REGION Network 11: External containerstation
         ON    "DB702_Tank_Value".Tank[1].With_ContainerStation;
         O     "DB009_Faults".Faults_Reset_FKT_M1;
         R     "DB822_Error_Tank".InterfaceContainer.FLT_SupplyContainerstation;
         R     "DB822_Error_Tank".InterfaceContainer.FLT_containerstation;
         R     "DB822_Error_Tank".InterfaceContainer.FLT_containerNotReady_C1;
   //-----
         AN    "Container_FaultSupply";
         A     "DB702_Tank_Value".Tank[1].With_ContainerStation;
         AN    "DB822_Error_Tank".InterfaceContainer.FLT_SupplyContainerstation;
         S     "DB822_Error_Tank".InterfaceContainer.FLT_SupplyContainerstation;
         S     "DB009_Faults".Faultschanging_M1;
   //---
   //      U     "Container_Faulty"
   //      U     "DB702_Tank_Value".Tank[1].With_ContainerStation
   //      UN    "DB822_Error_Tank".InterfaceContainer.FLT_containerstation
   //      S     "DB822_Error_Tank".InterfaceContainer.FLT_containerstation
   //      S     "DB009_Faults".Faultschanging_M1
   //---
         A     "ES_Container_C1";
         A     "DB702_Tank_Value".Tank[1].With_ContainerStation;
         =     "DB822_Error_Tank".InterfaceContainer.MSG_EScontainerstation;
   //---
         AN    "Container_Ready_C1";
         A     "DB702_Tank_Value".Tank[1].With_ContainerStation;
         A     "DB612_Tank_State".Tank[1].Switch_Refilling_ON_OFF;
         A     "DB619_State_MPart".Operationmode[1].Controllvoltage;
         AN    "DB822_Error_Tank".InterfaceContainer.FLT_containerNotReady_C1;
         S     "DB822_Error_Tank".InterfaceContainer.FLT_containerNotReady_C1;
         S     "DB009_Faults".Faultschanging_M1;
   //---
         AN    "Container_Ready_C1";
         A     "DB702_Tank_Value".Tank[1].With_ContainerStation;
         A     "DB619_State_MPart".Operationmode[1].Controllvoltage;
         A     "DB612_Tank_State".Tank[1].Switch_Refilling_ON_OFF;
         AN    "DB822_Error_Tank".InterfaceContainer.FLT_containerNotReady_C1;
         =     "DB822_Error_Tank".InterfaceContainer.MSG_containerNotReady_C1;
   //---
         O     "DB822_Error_Tank".InterfaceContainer.FLT_SupplyContainerstation;
         O     "DB822_Error_Tank".InterfaceContainer.FLT_containerstation;
         O     "DB822_Error_Tank".InterfaceContainer.FLT_containerNotReady_C1;
         S     "DB009_Faults".Faults_FKT_Grp_3_M1;
   //---
END_REGION

REGION Network 12: A fault exists
         O     "DB612_Tank_State".Tank[1].Fault_Exist;
         O     "DB612_Tank_State".Agitator[1].FLT_Exist;
         O     "DB612_Tank_State".AgitatorBarell[1].FLT_Exist;
         O     "DB612_Tank_State".Vacuum[1].FLT_PVacuum;
         O     "DB612_Tank_State".CirculationPump[1].FaultExist;
         O     "DB612_Tank_State".ControllerTankTemp[1].Fault_Exist;
         O     "DB612_Tank_State".ControllerTankJacketHeater[1].Fault_Exist;
         O     "DB612_Tank_State".ControllerBarellTemp[1].Fault_Exist;
   //---
         O     "DB822_Error_Tank".InterfaceContainer.FLT_SupplyContainerstation;
         O     "DB822_Error_Tank".InterfaceContainer.FLT_containerstation;
         O     "DB822_Error_Tank".InterfaceContainer.FLT_containerNotReady_C1;
   //---
         =     "DB612_Tank_State".FaultExists[1];
END_REGION
END_FUNCTION_BLOCK

FUNCTION_BLOCK "FB102_Common_Aggregates_C2"   // FB102, STL
TITLE = Agitators,Tanks, Refilling, tempering
{ S7_Optimized_Access := 'FALSE' }
AUTHOR : KT242
VERSION : 0.1
// Common aggregates
   VAR_TEMP
      DINT_dummy : Real;
      CompUsedForShot : Array[1..16] of Bool;
      Dummy : Bool;
      MH_open : Bool;
      K_Tanklager : Bool;
      Valid : Bool;
      Temp_Vacuum_active : Bool;
      Temp_Cooling : Bool;
      Temp_Filling_Enable : Bool;
      Temp_StartExtern : Bool;
      Temp_WithFillingPump : Bool;
      Temp_FillingPumpActive : Bool;
      Temp_SwitchONTemp : Bool;
      Temp_EnableTempering : Bool;
      Temp_RequestFillAuto : Bool;
      HF_Pulse_alarm : Bool;
      Temp_RetVal_SFC14 : Word;
      Temp_RetVal_SFC15 : Word;
      Temp_SetValue_TG : Int;
      Temp_Refilling_Barrel : Bool;
      Temp_Filling_Valve : Bool;
   END_VAR
BEGIN

REGION Network 1: Toggle bit, if refilling over barrel station is activated
   // Copy Control bits for module to local area
         L;
         LAR1;
         L     "DB619_State_MPart".ShotMa[1].ShotData.Comp_at_Shot;
         L     "DB619_State_MPart".ShotMa[2].ShotData.Comp_at_Shot;
         OD;
         CAW;
         T     LW [ AR1 , P#0.0 ];

         A     "DB612_Tank_State".Tank[2].Switch_Refilling_from_Barrel_ON_OFF;
         =     #Temp_Refilling_Barrel;
END_REGION

REGION Network 2: Signal a mixinghead opens
         O     "DB619_State_MPart".Mixinghead[1].Shotcounter."01";
         O     "DB619_State_MPart".Mixinghead[1].Shotcounter."02";
         O     "DB619_State_MPart".Mixinghead[1].Shotcounter."03";
         O     "DB619_State_MPart".Mixinghead[1].Shotcounter."04";
         O     "DB619_State_MPart".Mixinghead[1].Shotcounter."05";
         O     "DB619_State_MPart".Mixinghead[1].Shotcounter."06";
         O     "DB619_State_MPart".Mixinghead[1].Shotcounter."07";
         O     "DB619_State_MPart".Mixinghead[1].Shotcounter."08";
         O     "DB619_State_MPart".Mixinghead[1].Shotcounter."09";
         O     "DB619_State_MPart".Mixinghead[1].Shotcounter."10";
         O     "DB619_State_MPart".Mixinghead[1].Shotcounter."11";
         O     "DB619_State_MPart".Mixinghead[1].Shotcounter."12";
         O     "DB619_State_MPart".Mixinghead[1].Shotcounter."13";
         O     "DB619_State_MPart".Mixinghead[1].Shotcounter."14";
         O     "DB619_State_MPart".Mixinghead[1].Shotcounter."15";
         O     "DB619_State_MPart".Mixinghead[1].Shotcounter."16";
         A     #CompUsedForShot[2];
         =     #MH_open;
END_REGION

REGION Network 3: Filling level
         CALL  "FC920_PV_Calc_Act_Value"
         ( IN_Act_Value_read := "DB702_Tank_Value".Tank[2].With_Level_Probe,
           IN_Act_Value_ext  := FALSE,
           IN_Ext_Value      := #DINT_dummy,
           IN_Read_Double    := FALSE,
           IN_FLT_Needful    := TRUE,
           IN_FLT_Reset      := "DB009_Faults".Faults_Reset_FKT_M1,
           IO_Any_ArrayPV    := "DB602_PV_Tank".Tank[2].Level,
           IO_Fault_Sensor   := "DB822_Error_Tank".Refilling_Tank[2].FLT_LevelSensor_broken_wire,
           IO_New_Fault      := "DB009_Faults".Faultschanging_M1,
           IO_FLT_Level_3    := "DB009_Faults".Faults_FKT_Grp_3_M1
         );
   //-----
         AN    "DB702_Tank_Value".Tank[2].DrainTank;
         R     "DB612_Tank_State".Tank[2].Switch_DrainTank_ON_OFF;
   //-----
         CALL  "FC104_FillingSignals"
         ( Tank_exist           := "DB702_Tank_Value".Tank[1].Existing,
           Actual_Level_Value   := "DB602_PV_Tank".Tank[2].Level.PV_ActV.Value,
           IN_With_Level_Probe  := "DB702_Tank_Value".Tank[2].With_Level_Probe,
           IN_With_Triptray     := "DB702_Tank_Value".Tank[2].With_Triptray,
           IN_FLT_Level_Probe   := "DB822_Error_Tank".Refilling_Tank[2].FLT_LevelSensor_broken_wire,
           IN_Max_Level         := "L_DT_max_C2",
           IN_Stop_Fill_Level   := "L_Tank_stop_C2",
           IN_Start_Fill_Level  := "L_Tank_start_C2",
           IN_Min_Level         := "L_Tank_min_C2",
           IN_Triptray          := "L_DripTray_C2",
           IN_DrainTank         := "DB612_Tank_State".Tank[2].Switch_DrainTank_ON_OFF,
           OUT_PreWarnMinLevel  := "DB612_Tank_State".Tank[2].PreWarning_Min_Level,
           OUT_Max_Level        := "DB612_Tank_State".Tank[2].Max_Level,
           OUT_Stop_Fill_Level  := "DB612_Tank_State".Tank[2].Stop_Level_Filling,
           OUT_Start_Fill_Level := "DB612_Tank_State".Tank[2].Start_Level_Filling,
           OUT_Min_Level        := "DB612_Tank_State".Tank[2].Min_Level,
           OUT_Enable_Agitator  := "DB612_Tank_State".Tank[2].Enable_Agitator,
           OUT_Triptray         := "DB612_Tank_State".Tank[2].LevelTriptray,
           IO_TankLevelPar      := "DB702_Tank_Value".Tank[2].TankLevel
         );
   //-----
END_REGION

REGION Network 4: GBE
   //      CALL  "FC920_PV_Calc_Act_Value"
   //         IN_Act_Value_read :="DB702_Tank_Value".Tank[2].With_Nucleation
   //         IN_Act_Value_ext  :=FALSE
   //         IN_Ext_Value      :=#DINT_dummy
   //         IN_Read_Double    :=FALSE
   //         IN_FLT_Needful    :=TRUE
   //         IN_FLT_Reset      :="DB009_Faults".Faults_Reset_FKT_M1
   //         IO_Any_ArrayPV    :="DB602_PV_Tank".Tank[2].Nucleation
   //         IO_Fault_Sensor   :="DB822_Error_Tank".Refilling_Tank[2].FLT_NucleationSensor_broken_wire
   //         IO_New_Fault      :="DB009_Faults".Faultschanging_M1
   //         IO_FLT_Level_3    :="DB009_Faults".Faults_FKT_Grp_3_M1
   //-----
   //      O     "DB009_Faults".Faults_Reset_FKT_M1
   //      O     "DB702_Tank_Value".Tank[2].With_Nucleation
   //      R     "DB822_Error_Tank".Refilling_Tank[2].FLT_supply_nucleation
   //      R     "DB822_Error_Tank".Refilling_Tank[2].FLT_nucleation
   //-
   //      UN    "F_GBE_C2"
   //      U     "DB702_Tank_Value".Tank[2].With_Nucleation
   //      UN    "DB822_Error_Tank".Refilling_Tank[2].FLT_supply_nucleation
   //      S     "DB009_Faults".Faultschanging_M1
   //      S     "DB822_Error_Tank".Refilling_Tank[2].FLT_supply_nucleation
   //-
   //      U     "F_GBE_Faulty_C2"
   //      U     "DB702_Tank_Value".Tank[2].With_Nucleation
   //      UN    "DB822_Error_Tank".Refilling_Tank[2].FLT_nucleation
   //      S     "DB009_Faults".Faultschanging_M1
   //      S     "DB822_Error_Tank".Refilling_Tank[2].FLT_nucleation
   //-
   //      O     "DB822_Error_Tank".Refilling_Tank[2].FLT_nucleation
   //      O     "DB822_Error_Tank".Refilling_Tank[2].FLT_supply_nucleation
   //      S     "DB009_Faults".Faults_FKT_Grp_3_M1
   //-----
END_REGION

REGION Network 5: Filling daytank
   ///----
         AN    "DB822_Error_Tank".FeedPump[2].FLT_Dryrunsafety;
         AN    "DB822_Error_Tank".FeedPump[2].FLT_Motorprotection;
         AN    "DB822_Error_Tank".FeedPump[2].FLT_No_Barrel;
         A(;
         ON    "DB702_Tank_Value".Tank[2].With_ContainerStation;
         O     "Container_Ready_C2";
         );
         A     "DB619_State_MPart".Operationmode[1].valid;
         =     #Temp_Filling_Enable;
   //-----
         A     "Container_Fillpump_run_C2";
         =     #Temp_FillingPumpActive;
   //-----
         A     "DB702_Tank_Value".Tank[2].With_ContainerStation;
         =     #Temp_WithFillingPump;
   //-----
         CALL  "FC102_Refilling"
         ( IN_Selected             := "DB702_Tank_Value".Tank[2].Existing,
           IN_ReleaseRefilling     := #Temp_Filling_Enable,
           IN_FillingPumpActive    := #Temp_FillingPumpActive,
           IN_WithFillingPump      := #Temp_WithFillingPump,
           IN_RecircWeekend        := "DB619_State_MPart".Recirculation[1].Weekendswitching,
           IN_FoamingCycleActive   := "DB619_State_MPart".Cycle[1].running,
           IN_PistonActive         := FALSE,
           IN_MH_is_open           := #MH_open,
           IN_ResetFault           := "DB009_Faults".Faults_Reset_FKT_M1,
           IN_MaxLevelTriptray     := "DB612_Tank_State".Tank[2].LevelTriptray,
           IN_PumpDeselected       := "DB753_MeteringPump".Pump[2].PumpDeselected,
           IN_SetAmountShots       := "DB702_Tank_Value".Tank[2].NoShotFilling,
           IN_PreAgitatingTime     := "DB702_Tank_Value".Tank[2].PreAgitatingTime,
           IN_FillingTimeContr     := "DB702_Tank_Value".Tank[2].FillingTimeControl,
           IN_TimeTillFillingStart := "DB702_Tank_Value".Tank[2].TimeToStartFilling,
           IN_Timer_Refilling      := "TM_Refilling_02",
           OUT_V_Preagitating      := #Dummy,
           OUT_V_Refilling         := #Temp_Filling_Valve,  //"V_ChargingTank_C2"
           OUT_R_Tankstorage       := #K_Tanklager,
           IO_Status               := "DB612_Tank_State".Tank[2],
           IO_NewFault             := "DB009_Faults".Faultschanging_M1,
           IO_FaultLevel_1         := "DB009_Faults".Faults_FKT_Grp_1_M1,
           IO_FaultLevel_2         := "DB009_Faults".Faults_FKT_Grp_2_M1,
           IO_FaultLevel_3         := "DB009_Faults".Faults_FKT_Grp_3_M1,
           IO_Fault                := "DB822_Error_Tank".Refilling_Tank[2]
         );
   //-----
         A     #Temp_Refilling_Barrel;
         JC    BarrelFill;
         R     "K_Filling_Tank_C2_TL";
         R     "V_ChargingTank_C2_2";

         A     #K_Tanklager;
         A     #Temp_Filling_Valve;
         =     "K_Filling_Tank_C2";
         =     "V_ChargingTank_C2";
         =     "V_Barrel_C2";
         =     "C_Start_Refill_ISO_ON";

         JU    NoBarrelFill;

   BarrelFill:R     "K_Filling_Tank_C2";
         R     "V_ChargingTank_C2";

         A     #K_Tanklager;
         A     #Temp_Filling_Valve;
         =     "K_Filling_Tank_C2_TL";
         =     "V_ChargingTank_C2_2";
         =     "V_Barrel_C2";
         =     "C_Start_Refill_ISO_ON";


   //-----
END_REGION

REGION Network 6: Agitator daytank
   //-----
   // Das Befüllen soll das Rührwerk nur im Auto ansteuern
   NoBarrelFill:A     "DB612_Tank_State".Tank[2].Fillingtime_runs;
         A     "DB619_State_MPart".Operationmode[1].Auto;
         =     #Temp_RequestFillAuto;

         CALL  "FC121_Aggitator"
         ( IN_Release               := "DB619_State_MPart".Operationmode[1].valid,
           IN_ControlVoltage        := "DB619_State_MPart".Operationmode[1].Controllvoltage,
           IN_Reset_fault           := "DB009_Faults".Faults_Reset_FKT_M1,
           IN_Request_Filling       := #Temp_RequestFillAuto,  //"DB612_Tank_State".Tank[2].Fillingtime_runs
           IN_Request_Feed          := 0,
           IN_Request_Cooling       := "DB612_Tank_State".ControllerTankTemp[2].CoolingActive,
           IN_Request_Heating       := "DB612_Tank_State".ControllerTankTemp[2].HeatingActive,
           IN_Fault_Motorprotection := "F_Agitator_C2",
           IN_FaultFreqConverter    := "F_FC_Agitator_C2",
           IN_MaxLevelTray          := "DB612_Tank_State".Tank[2].LevelTriptray,
           IN_EnableLevel           := "DB612_Tank_State".Tank[2].Enable_Agitator,
           IN_TimerDrive            := "TM1_Agitator_02",
           IN_TimerStartUpFConv     := "TM2_Agitator_02",
           IN_Values                := "DB702_Tank_Value".Tank[2].Agitator,
           OUT_MainsContactor       := "M_Agitator_C2",
           OUT_Release_FConverter   := "M_FU_Start_RW_K2",
           IO_Status                := "DB612_Tank_State".Agitator[2],
           IO_NewFault              := "DB009_Faults".Faultschanging_M1,
           IO_FaultLevel_3          := "DB009_Faults".Faults_FKT_Grp_3_M1,
           IO_Faults                := "DB822_Error_Tank".Agitator[2]
         );
   //-----
END_REGION

REGION Network 7: Tempering Tank
         A     "DB009_Faults".Faults_Reset_FKT_M1;
         R     "DB822_Error_Tank".ControllerTankTemp[2].Fuse_TemperingUnit;
   //-
         AN    "F_Temperiergeraet_C2";
         A     "DB702_Tank_Value".Tank[2].With_Tempering_TempGeraet;
         AN    "DB822_Error_Tank".ControllerTankTemp[2].Fuse_TemperingUnit;
         S     "DB009_Faults".Faultschanging_M1;
         S     "DB822_Error_Tank".ControllerTankTemp[2].Fuse_TemperingUnit;
   //-
         A     "DB822_Error_Tank".ControllerTankTemp[2].Fuse_TemperingUnit;
         S     "DB009_Faults".Faults_FKT_Grp_3_M1;
   //-
         CALL  "FC920_PV_Calc_Act_Value"
         ( IN_Act_Value_read := TRUE,
           IN_Act_Value_ext  := FALSE,
           IN_Ext_Value      := #DINT_dummy,
           IN_Read_Double    := FALSE,
           IN_FLT_Needful    := TRUE,
           IN_FLT_Reset      := "DB009_Faults".Faults_Reset_FKT_M1,
           IO_Any_ArrayPV    := "DB602_PV_Tank".Tank[2].Temp,
           IO_Fault_Sensor   := "DB822_Error_Tank".ControllerTankTemp[2].Sensor_FLT_broken_wire,
           IO_New_Fault      := "DB009_Faults".Faultschanging_M1,
           IO_FLT_Level_3    := "DB009_Faults".Faults_FKT_Grp_3_M1
         );
   //-----
         CALL  "FC916_PV_Limits"
         ( IN_Tolerance_Test     := TRUE,
           IN_Reset_Fault        := "DB009_Faults".Faults_Reset_FKT_M1,
           IO_Any_ArrayPV        := "DB602_PV_Tank".Tank[2].Temp,
           IO_Fault_Warn_upperL  := "DB822_Error_Tank".ControllerTankTemp[2].Warning_limit_plus,
           IO_Fault_Warn_lowerL  := "DB822_Error_Tank".ControllerTankTemp[2].Warning_limit_minus,
           IO_Fault_Alarm_upperL := "DB822_Error_Tank".ControllerTankTemp[2].Alarm_limit_plus,
           IO_Fault_Alarm_lowerL := "DB822_Error_Tank".ControllerTankTemp[2].Alarm_limit_minus,
           IO_New_Fault          := "DB009_Faults".Faultschanging_M1,
           IO_Fault_Level_1      := "DB009_Faults".Faults_FKT_Grp_2_M1,
           IO_Fault_Level_2      := #Dummy,  //"DB009_Faults".Faults_FKT_Grp_2_M1
           IO_Fault_Level_3      := "DB009_Faults".Faults_FKT_Grp_3_M1
         );
   //-----
   //---------------------------------------------
   //  Controller temperature tank Iso
   //---------------------------------------------
         O     "DB702_Tank_Value".Tank[2].With_Tempering_VKaltwasser;
         O     "DB702_Tank_Value".Tank[2].With_Tempering_Heizung;
         =     #Temp_EnableTempering;
   //---
         CALL  "FC105_Tempering"
         ( IN_Exist                := #Temp_EnableTempering,
           IN_Release              := "DB619_State_MPart".Operationmode[1].valid,
           IN_Stop_Tempering       := FALSE,
           IN_F_Fuse               := "F_Heating",
           IN_F_Limit              := FALSE,
           IN_FLT_Ackn             := "DB009_Faults".Faults_Reset_FKT_M1,
           IN_CoolingRequested     := TRUE,
           IN_HeatingRequested     := "DB702_Tank_Value".Tank[2].With_Tempering_Heizung,
           IN_actual_Temp          := "DB602_PV_Tank".Tank[2].Temp.PV_ActV.Value,
           IN_set_Temp             := "DB602_PV_Tank".Tank[2].Temp.PV_SetV.Value,
           Out_act_cooling         := #Temp_Cooling,
           Out_act_request_cooling := #Dummy,
           Out_act_heating         := "K_HeatingTank_C2",
           Out_act_request_heating := #Dummy,
           IO_StateCtrl1           := "DB612_Tank_State".ControllerTankTemp[2],
           IO_ValueCtrl1           := "DB702_Tank_Value".Pt2_Controller[2],
           IO_FaultsCtrl1          := "DB822_Error_Tank".ControllerTankTemp[2],
           IO_NewFault             := "DB009_Faults".Faultschanging_M1,
           IO_FaultLevel_3         := "DB009_Faults".Faults_FKT_Grp_3_M1
         );
   //-----
         A     "DB619_State_MPart".Machine[1].Metering."02";
         A     "DB702_Tank_Value".Tank[2].With_Tempering_WTRL;
         A     #Temp_Cooling;
         O(;
         A     "DB613_Komponent_State".HeatexchangerLP[2].CoolingActive;
         A     "DB619_State_MPart".Machine[1].Metering."02";
         A     "DB753_MeteringPump".Pump[2].WithLPHeatExchanger;
         );
         =     "V_Heatexchanger_C2";
   //-----
         ON    "DB619_State_MPart".Machine[1].Metering."02";
         ON    "DB702_Tank_Value".Tank[2].With_Tempering_WTRL;
         A     #Temp_Cooling;
         =     "V_Coolingwater_C2";
   //-----

   // Tempering device gets/sets temperature values with multiplier of 10.
         CALL  CONVERTTO
         ( IN      := "DB602_PV_Tank".Tank[2].Temp.PV_SetV.Value,
           Ret_Val := #Temp_SetValue_TG
         );

         L     #Temp_SetValue_TG;
         L     10;
         *I;
         T     #Temp_SetValue_TG;

         A     "Flag_00_500_Hertz";
         FP    "HF_pulse_alarm_GWK2";
         =     #HF_Pulse_alarm;

   //     CALL  "GWK_PB_TecoCS(CW)e"
   //         IN_With_tempering_unit :="DB702_Tank_Value".Tank[2].With_Tempering_TempGeraet
   //         IN_Flag_alarm          :=#HF_Pulse_alarm
   //         IN_Adr                 :="gwk_temp2~gwk_KRPRO_V6_2_1"
   //         IN_Sl_Akt              :=1
   //         IN_TL_KomF             :=1
   //         IN_On                  :="DB612_Tank_State".ControllerTankTemp[2].Switch_Temp_ON_OFF
   //         IN_Release             :="DB619_State_MPart".Operationmode[1].valid//"DB10_State_MC1".Operating_mode.valid
   //         IN_Weekendmode         :=FALSE
   //         IN_Fault_quit          :="DB009_Faults".Faults_Reset_FKT_M1
   //         IN_Fuse                :="F_Temperiergeraet_C2"
   //         IN_Setvalue            :=#Temp_SetValue_TG
   //         IN_Setvalue_weekend    :=#Temp_SetValue_TG
   //         IN_Actvalue_tool       :="DB602_PV_Tank".Tank[2].Temp.PV_ActV.Value
   //         RetVal_SFC14           :=#Temp_RetVal_SFC14
   //         RetVal_SFC15           :=#Temp_RetVal_SFC15
   //         PBData                 :="DB905_GWK".teco_cs_cw_e[2]
   //         State                  :="DB905_GWK".State[2]
END_REGION

REGION Network 8: Filling pump
         A     "DB009_Faults".Faults_Reset_FKT_M1;
         R     "DB822_Error_Tank".FeedPump[2].FLT_Dryrunsafety;
         R     "DB822_Error_Tank".FeedPump[2].FLT_Motorprotection;
         R     "DB822_Error_Tank".FeedPump[2].FLT_No_Barrel;
   //----- Störung Trockenlauf Befüllung
         A(;
         O     "K_Filling_Tank_C2";
         O     "K_Filling_Tank_C2_TL";
         );
         A     "DB702_Tank_Value".Tank[2].With_Filling_DryRun;
         L     s5t#5s;
         SD    "TM_Tank_Delay_DryRun_FeedPump_C2";
   //---
         A     "TM_Tank_Delay_DryRun_FeedPump_C2";
         AN    "S_DryRun_Feed_C2";
         AN    "DB822_Error_Tank".FeedPump[2].FLT_Dryrunsafety;
         S     "DB822_Error_Tank".FeedPump[2].FLT_Dryrunsafety;
         S     "DB009_Faults".Faults_FKT_Grp_3_M1;
         S     "DB009_Faults".Faultschanging_M1;
   //----- Störung Motorschutz Füllpumpe
         A     "F_FeedPump_C2";
         A     "DB702_Tank_Value".Tank[2].With_Filling_Pump;
         AN    "DB822_Error_Tank".FeedPump[2].FLT_Motorprotection;
         S     "DB822_Error_Tank".FeedPump[2].FLT_Motorprotection;
         S     "DB009_Faults".Faults_FKT_Grp_3_M1;
         S     "DB009_Faults".Faultschanging_M1;
   //----- Störung Kein Fass vorhanden aber Befüllung angewählt
   //    U     "K_Filling_Tank_C2"
   //    UN    "S_BarrelDetection_C2"
   //    UN    "DB822_Error_Tank".FeedPump[2].FLT_No_Barrel
   //    S     "DB822_Error_Tank".FeedPump[2].FLT_No_Barrel
   //    S     "DB009_Faults".Faults_FKT_Grp_3_M1
   //    S     "DB009_Faults".Faultschanging_M1
   //----- Meldung Kein Fass vorhanden
   //    UN    "S_BarrelDetection_C2"
   //    UN    "DB822_Error_Tank".FeedPump[2].FLT_No_Barrel
         CLR;
         =     "DB822_Error_Tank".FeedPump[2].Mes_No_Barrel;
   //-----
         AN    "DB822_Error_Tank".FeedPump[2].FLT_No_Barrel;
         AN    "DB822_Error_Tank".FeedPump[2].Mes_No_Barrel;
         AN    "DB822_Error_Tank".FeedPump[2].FLT_Dryrunsafety;
         AN    "DB822_Error_Tank".FeedPump[2].FLT_Motorprotection;
         A(;
         O     "K_Filling_Tank_C2";
         O     "K_Filling_Tank_C2_TL";
         );
         =     "M_FeedPump_C2";
   //-----
END_REGION

REGION Network 9: Vacuum daytank
         CALL  "FC106_Vacuum"
         ( IN_Release           := "DB619_State_MPart".Operationmode[1].valid,
           IN_P_Vacuum          := "P_Vacuum_C2",
           IN_Timer_delay_Lock  := "TM_Vac2DelayLock",
           IN_Timer_delay_Pumpe := "TM_Vac2DelayPump",
           OUT_V_Lock_Vacuum    := "V_PressureVacuum_C2",
           OUT_V_Pump_Vacuum    := "V_PumpVacuum_C2",
           OUT_H_Vacuum_active  := #Temp_Vacuum_active,
           IO_Status            := "DB612_Tank_State".Vacuum[2]
         );
   //-----
END_REGION

REGION Network 10: High pressure heatexchanger
   // ------------------------------------------------------
   // Heatexchanger K1
   // ------------------------------------------------------
   //      CALL  "FC920_PV_Calc_Act_Value"
   //         IN_Act_Value_read :=TRUE
   //         IN_Act_Value_ext  :=FALSE
   //         IN_Ext_Value      :=#DINT_dummy
   //         IN_Read_Double    :=FALSE
   //         IN_FLT_Reset      :="DB009_Faults".Faults_Reset_FKT_M1
   //         IO_Any_ArrayPV    :="DB603_PV_Tempering".Tempering_Heatexchanger[1].Temperature_1
   //         IO_Fault_Sensor   :="DB810_Error_general".Temperature_Heatexchange[1].Sensor_FLT_broken_wire
   //         IO_New_Fault      :="DB009_Faults".Faultschanging_M1
   //         IO_FLT_Level_3    :="DB009_Faults".Faults_FKT_Grp_3_M1
   //-------------------------------------------------------
   // Check limits temperature C1 Heatexchanger
   //-------------------------------------------------------
   //      CALL  "FC916_PV_Limits"
   //         IN_Tolerance_Test     :="DB610_State_MPart".Operationmode_Ma[1].Controllvoltage
   //         IN_Reset_Fault        :="DB121_PUC08_PLC_State".IN_PUC.Status_M1.FLT_quit_from_PLC
   //         IO_Any_ArrayPV        :="DB603_PV_Tempering".Tempering_Heatexchanger[1].Temperature_1
   //         IO_Fault_Warn_upperL  :="DB810_Error_general".Temperature_Heatexchange[1].Warning_limit_plus
   //         IO_Fault_Warn_lowerL  :="DB810_Error_general".Temperature_Heatexchange[1].Warning_limit_minus
   //         IO_Fault_Alarm_upperL :="DB810_Error_general".Temperature_Heatexchange[1].Alarm_limit_plus
   //         IO_Fault_Alarm_lowerL :="DB810_Error_general".Temperature_Heatexchange[1].Alarm_limit_minus
   //         IO_New_Fault          :="DB009_Faults".Faultschanging_M1
   //         IO_Fault_Level_1      :="DB009_Faults".Faults_FKT_Grp_1_M1
   //         IO_Fault_Level_2      :="DB009_Faults".Faults_FKT_Grp_2_M1
   //         IO_Fault_Level_3      :="DB009_Faults".Faults_FKT_Grp_3_M1
   //
   //------------------------------------------------------------
   //  Controller temperature Headexchanger C1 pulse width control
   //------------------------------------------------------------
   //      U(
   //      L     "DB603_PV_Tempering".Tempering_Heatexchanger[1].Temperature_1.PV_Conf_ActV.ControllerType
   //      L     2
   //      ==I
   //      )
   //      U(
   //      L     "DB603_PV_Tempering".Tempering_Heatexchanger[1].Temperature_1.PV_Conf_ActV.ControllerNo
   //      L     0
   //      >I
   //      )
   //      SPBN  EHD1
   //
   //
   //      CALL  "FC151_ReadArrayToZero"
   //         Nr_Array   :="DB603_PV_Tempering".Tempering_Heatexchanger[1].Temperature_1.PV_Conf_ActV.ControllerNo
   //         LowerLimit :=1
   //         UpperLimit :=64
   //         Any_Cont   :="DB780_Para_PW-Control".PW_Controller[0]
   //
   //      L     "DB603_PV_Tempering".Tempering_Heatexchanger[1].Temperature_1.PV_ActV.Value
   //      L     10
   //      /D
   //      T     #Temp_HD_WT
   //
   //      L     "DB603_PV_Tempering".Tempering_Heatexchanger[1].Temperature_1.PV_SetV.Value
   //      L     10
   //      /D
   //      T     #Temp_SetValueTemp
   //
   //      L     "DB780_Para_PW-Control".PW_Controller[0].Max_Temp_Diff_Cooling
   //      L     10
   //      /D
   //      T     #Pulse_K1_MaxDelta_K
   //
   //      L     "DB780_Para_PW-Control".PW_Controller[0].Max_Temp_Diff_Heating
   //      L     10
   //      /D
   //      T     #Pulse_K1_MaxDelta_H
   //
   //      CALL  "FC56_TemPulse2"
   //         Trig              :="TriggerPulse"
   //         In_Sollwert       :=#Temp_SetValueTemp
   //         In_Istwert_Tank   :=#Temp_HD_WT
   //         In_Istwert_Return :=#Temp_HD_WT
   //         In_Wichtung       :="DB780_Para_PW-Control".PW_Controller[0].Weighting_Temp
   //         In_Regelstrecke   :="DB780_Para_PW-Control".PW_Controller[0].PLC_Control_Area
   //         In_MaxDelta_K     :=#Pulse_K1_MaxDelta_K
   //         In_MaxDelta_H     :=#Pulse_K1_MaxDelta_H
   //         Pulsezeit         :="HDTempPulseTime_K1"//"DB610_State_MPart".Controller[0].PulsTime
   //         Heating           :=#Dummy
   //         Cooling           :=#Temp_Cooling
   //
   //
   // Regelstrecke von PUC auf ms Format
   //      L     "DB780_Para_PW-Control".PW_Controller[0].PLC_Control_Area
   //      L     1000
   //      *D
   //      T     #Regelstrecke        // Zeitwert für Timer
   //
   // Regelstreckentimer ständig starten
   //      UN    "TriggerPulse"
   //      =     "StartDelayTimer"
   //
   //      CALL  TON , "DB55_Temp_HD_WT_MK1_K1"
   //         IN :="StartDelayTimer"
   //         PT :=#Regelstrecke
   //         Q  :="TriggerPulse"
   //         ET :=#Zeit_abgelaufen
   //
   // Kühlen  EIN
   //      U     #Temp_Cooling
   //      S     "HM_HDWT_MH1_K1_cool"
   //
   // Kühlen  AUS
   //      L     "HDTempPulseTime_K1"
   //      L     #Zeit_abgelaufen
   //      <D
   //      UN(
   //      L     "HDTempPulseTime_K1"
   //      L     #Regelstrecke
   //      >D
   //      )
   //      ON    "DB128_KeysSignals_B&R".T_BR_Key_ON[11]
   //      ON    "DB610_State_MPart".Operationmode_Ma[1].valid
   //      O     "DB810_Error_general".Temperature_Heatexchange[1].Sensor_FLT_broken_wire
   //      R     "HM_HDWT_MH1_K1_cool"
   //
   //      U     "HM_HDWT_MH1_K1_cool"
   //      U     "DB121_PUC08_PLC_State".IN_PUC.Metering._01
   //      =     #Dummy
   //      =     "V_HDWT_Kuehl_K1_M1"        // stromlos zu
   //      =     "V_HDWT_Bypass_K1_M1"       // stromlos offen
   //
   //EHD1: NOP 0
END_REGION

REGION Network 11: External containerstation
         ON    "DB702_Tank_Value".Tank[2].With_ContainerStation;
         O     "DB009_Faults".Faults_Reset_FKT_M1;
         R     "DB822_Error_Tank".InterfaceContainer.FLT_SupplyContainerstation;
         R     "DB822_Error_Tank".InterfaceContainer.FLT_containerstation;
         R     "DB822_Error_Tank".InterfaceContainer.FLT_containerNotReady_C2;
   //-----
         AN    "Container_FaultSupply";
         A     "DB702_Tank_Value".Tank[2].With_ContainerStation;
         AN    "DB822_Error_Tank".InterfaceContainer.FLT_SupplyContainerstation;
         S     "DB822_Error_Tank".InterfaceContainer.FLT_SupplyContainerstation;
         S     "DB009_Faults".Faultschanging_M1;
   //---
   //      U     "Container_Faulty"
   //      U     "DB702_Tank_Value".Tank[2].With_ContainerStation
   //      UN    "DB822_Error_Tank".InterfaceContainer.FLT_containerstation
   //      S     "DB822_Error_Tank".InterfaceContainer.FLT_containerstation
   //      S     "DB009_Faults".Faultschanging_M1
   //---
         A     "ES_Container_C1";
         A     "DB702_Tank_Value".Tank[2].With_ContainerStation;
         =     "DB822_Error_Tank".InterfaceContainer.MSG_EScontainerstation;
   //---
         AN    "Container_Ready_C2";
         A     "DB702_Tank_Value".Tank[2].With_ContainerStation;
         A     "DB612_Tank_State".Tank[2].Switch_Refilling_ON_OFF;
         A     "DB619_State_MPart".Operationmode[1].Controllvoltage;
         AN    "DB822_Error_Tank".InterfaceContainer.FLT_containerNotReady_C2;
         S     "DB822_Error_Tank".InterfaceContainer.FLT_containerNotReady_C2;
         S     "DB009_Faults".Faultschanging_M1;
   //---
         AN    "Container_Ready_C2";
         A     "DB702_Tank_Value".Tank[2].With_ContainerStation;
         A     "DB619_State_MPart".Operationmode[1].Controllvoltage;
         A     "DB612_Tank_State".Tank[2].Switch_Refilling_ON_OFF;
         AN    "DB822_Error_Tank".InterfaceContainer.FLT_containerNotReady_C2;
         =     "DB822_Error_Tank".InterfaceContainer.MSG_containerNotReady_C2;
   //---
         O     "DB822_Error_Tank".InterfaceContainer.FLT_SupplyContainerstation;
         O     "DB822_Error_Tank".InterfaceContainer.FLT_containerstation;
         O     "DB822_Error_Tank".InterfaceContainer.FLT_containerNotReady_C2;
         S     "DB009_Faults".Faults_FKT_Grp_3_M1;
   //-----
END_REGION

REGION Network 12: A fault exists
         O     "DB612_Tank_State".Tank[2].Fault_Exist;
         O     "DB612_Tank_State".Agitator[2].FLT_Exist;
         O     "DB612_Tank_State".AgitatorBarell[2].FLT_Exist;
         O     "DB612_Tank_State".Vacuum[2].FLT_PVacuum;
         O     "DB612_Tank_State".CirculationPump[2].FaultExist;
         O     "DB612_Tank_State".ControllerTankTemp[2].Fault_Exist;
         O     "DB612_Tank_State".ControllerTankJacketHeater[2].Fault_Exist;
         O     "DB612_Tank_State".ControllerBarellTemp[2].Fault_Exist;
   //---
         O     "DB822_Error_Tank".InterfaceContainer.FLT_SupplyContainerstation;
         O     "DB822_Error_Tank".InterfaceContainer.FLT_containerstation;
         O     "DB822_Error_Tank".InterfaceContainer.FLT_containerNotReady_C2;
   //---
         =     "DB612_Tank_State".FaultExists[2];
END_REGION
END_FUNCTION_BLOCK

FUNCTION_BLOCK "FB110_Interface_Prog_M1"   // FB110, STL
TITLE = Interface mould carrier, external plant, FIFO
{ S7_Optimized_Access := 'FALSE' }
AUTHOR : KT242
VERSION : 0.1
   VAR_TEMP
      Release_Foaming_1 : Bool;   // Allgemeine Freigabe zum Starten des Schäumzyklusses der Schnittstelle
      TempReleasInterface : Bool;   // Freigabe von der Schnittstelle zum Starten des Schäumzyklusses
      Start_Zyklus : Bool;   // Impuls zum Starten des Schäumzyklusses
      Start_Zyklus_Roboter : Bool;   // Impuls zum Starten des Roboterprogrammes
      Automatik_Stop_ist_Quitt : Bool;   // Das Signal Automatik- Stopp wurde quittert, Automatikbetrieb ist ok
      Freigabe_Eintrag_von_PUC : Bool;   // Die Freigabe zum Schaumeintrag des Roboter von dem Rechner steht an
      Dummy : Bool;   // Dummybit für nicht benötigte Bausteinparameter
      Imp_Testschuss : Bool;   // Impulsmerker für die Anforderung eines automatischen Testschusses
      Imp_Tuer_1_Roboter : Bool;   // Impulsmerker für das öffnen/ schließen der Schutztür zum Roboter
      HM_Tuer_Auf : Bool;   // Hilfsmerker für das öffnen der Schutztür zum Roboter
      HM_Tuer_Zu : Bool;   // Hilfsmerker für das schließen der Schutztür zum Roboter
      MK_Reinigung_sofort : Bool;   // Die Mischkopf- Reinigung soll nach diesem Programm gestartet werden
      H_MH_Panel : Bool;
      Temp_Stop : Bool;
      Temp_ProgNo_MK1_manual : Byte;   // Programmvorwahl für Handschuss
      Speicher_PRG_NR_Hand : Word;   // Speicher für Programmnummer in Hand 1 bis 99 Programme
      Release_Foaming : Bool;   // Allgemeine Freigabe zum Starten des Schäumzyklusses der Schnittstelle
      Release_from_IF : Bool;   // Freigabe von der Schnittstelle zum Starten des Schäumzyklusses
      Start_Foaming : Bool;   // Impuls zum Starten des Schäumzyklusses
      Release_Datatransfer_Rob : Bool;   // Freigabe für die Übertragung der Programmnummer an den Roboter
      Start_Datatransfer : Bool;   // Starten der Übertragung der Programmnummer an den Roboter
      Release_Rob_Move : Bool;   // Freigabe für die Bewegung des Roboters in die Form
      Start_Rob_Move : Bool;   // Impuls zum Starten der Bewegung des Roboters in die Form
      E_Stop_quitt : Bool;   // Das Signal Automatik- Stopp wurde quittert, Automatikbetrieb ist ok
      Release_Foam_from_PUC : Bool;   // Die Freigabe zum Schaumeintrag des Roboter von dem Rechner steht an
      Temp_Teachen : Bool;   // Impulsmerker zum anfahren der Position zum Teachen
      Dummy_1 : Bool;   // Dummy- Merker zum belegen nicht verwendeter Ausgänge
      Drop_Wobj : Bool;   // Ein schon Syncronisiertes Werkobjekt wird gelöscht
      Release_WaitWobj : Bool;   // Freigabe zum aufsyncronisieren eines Werkobjektes
      EM_StartMoveHomepos : Bool;   // Freigabe für eine automatische fahrt in die Homeposition
      PointerDB : DWord;
      Automatik_Stop_ist_Qu_1 : Bool;
      Temp_Frg : Bool;
      Spuelmittel_Ein : Bool;
      V_Trocknen_Reiniger : Bool;
      V_Kreislauf_Reiniger : Bool;
      V_Spuelen_Reiniger : Bool;
      K_Heizung_Reiniger : Bool;
      V_Dichtung_Reiniger : Bool;
      Imp_Tuer_2_Roboter : Bool;
      HM_Tuer_2_Auf : Bool;   // Hilfsmerker für das öffnen der Schutztür zum Roboter
      HM_Tuer_2_Zu : Bool;   // Hilfsmerker für das schließen der Schutztür zum Roboter
      Temp_ProgNo_MK2_manual : Byte;
      Temp_Start_MK1 : Bool;
      Temp_Stop_MK1 : Bool;
      Temp_Manual_MK1 : Bool;
      Temp_Lamp_MK1 : Bool;
      Temp_Einer : Byte;
      Temp_Imp_Tuer_Roboter : Bool;
      Temp_OperateWithRobot : Bool;
      Temp_PrgNrDeselect : Bool;
      Temp_ProgNo_MK3_manual : Byte;
      Temp_ProgNo_MK4_manual : Byte;
      Temp_ProgNo_MK5_manual : Byte;
      Temp_ProgNo_MK6_manual : Byte;
      Temp_ProgNo_MK7_manual : Byte;
      Temp_ProgNo_MK8_manual : Byte;
      Temp_ProgNo_MK9_manual : Byte;
      Temp_ProgNo_MK10_manual : Byte;
   END_VAR
BEGIN

REGION Network 1: FIFO saves number of interface
         CALL  "FC111_FIFO"
         ( IN_Amount_Interfaces := "DB790_PlantParameter".AmountToolStation,
           IN_Register          := "DB110_Interf_Program_M1".Putin_FIFOlist,
           IN_Reset_List        := "Flag_Erster_SPS_Zyklus",
           IN_StartAdr          := "DB110_Interf_Program_M1".FIFO.FIFO_01.%B1,
           IN_DataBlock         := "DB110_Interf_Program_M1",
           IO_FIRST             := "DB110_Interf_Program_M1".FIRST,
           IO_SECOND            := "DB110_Interf_Program_M1".SECOND,
           IO_FlagNewPos        := "DB110_Interf_Program_M1".Bits.Ageflag
         );
END_REGION

REGION Network 2: Interface to external plant

         AN    "DB704_MH_Value".Mixinghead[1].Conf_IntWithPlantInerface;
         JC    NoInterfaceMH1;

         A     "DB619_State_MPart".Operationmode[1].Auto;
         A     "DB704_MH_Value".Mixinghead[1].Conf_IntWithPlantInerface;
         =     #TempReleasInterface;

         O(;
         A(;
         O     "DB614_MH_State".InertingMH[1].OK;
         O     "DB614_MH_State".InertingMH[1].Start_PressurizeTimeRuns;
         );
         FP    "DB614_MH_State".InertingMH[1].Reserve47;
         );
         A     "DB704_MH_Value".MH_Inerting[1].with_inert_over_MH;
         O(;
         A     "DB110_Interf_Program_M1".Signals_ExPlant[1].Strobe;
         AN    "DB704_MH_Value".MH_Inerting[1].with_inert_over_MH;
         );
         A     #TempReleasInterface;
         =     #Start_Zyklus;

         CALL  "FC114_IF_externalPlant"
         ( IN_Release               := #TempReleasInterface,
           IN_use_Inv_Program       := FALSE,
           IN_use_Parity_Bit        := FALSE,
           IN_Reset_fault_Fkt       := "DB009_Faults".Faults_Reset_FKT_M1,
           IN_Stop_MH_OpPanel       := "DB123_MH_IO_Signals".MH[1].IN.MH_Stop,
           IN_Operationmode_Operate := "DB619_State_MPart".Operationmode[1].Operation,
           IN_MH_panel_automatic    := "DB123_MH_IO_Signals".MH[1].IN.MH_Auto_Mode,
           IN_FCycleRelease_extern  := TRUE,
           IN_FCycle_release        := "DB619_State_MPart".Cycle[1].Release,
           IN_FCycle_running        := "DB619_State_MPart".Cycle[1].running,
           IN_FCycle_Shotrelease    := "DB619_State_MPart".Cycle[1].Shotrelease,
           IN_FCycle_Shot_running   := "DB619_State_MPart".Cycle[1].ShotRuns,
           IN_FCycle_Pulse_Shotend  := "DB619_State_MPart".Cycle[1].PulsShotend,
           IN_FCycle_Pulse_End      := "DB619_State_MPart".Cycle[1].PulseCycleEnd,
           IN_ExtPlant_OK           := "DB110_Interf_Program_M1".Signals_ExPlant[1].ExtP_OK,
           IN_Strobe_or_Start       := #Start_Zyklus,  //"DB110_Interf_Program_M1".Signals_ExPlant[1].Strobe
           IN_StrobeINV_or_Parity   := FALSE,
           IN_Start_Shot            := "DB110_Interf_Program_M1".Signals_ExPlant[1].MH_open,
           IN_CP_forward            := "DB110_Interf_Program_M1".Signals_ExPlant[1].CP_forward,
           IN_ProgNo_ExtPlant       := "DB110_Interf_Program_M1".Signals_ExPlant[1].PrgNo,
           IN_maxAmount_ProgNo      := 255,
           OUT_PU_OK                := "DB110_Interf_Program_M1".Signals_ExPlant[1].PU_OK,
           OUT_Strobe_quit          := "DB110_Interf_Program_M1".Signals_ExPlant[1].Strobe_quitt,
           OUT_FCycle_running       := "DB110_Interf_Program_M1".Signals_ExPlant[1].cycle_run,
           OUT_ReadyForFoaming      := "DB110_Interf_Program_M1".Signals_ExPlant[1].ready_for_shot,
           OUT_FoamingActive        := "DB110_Interf_Program_M1".Signals_ExPlant[1].shot_run,
           OUT_FoamingEnd           := "DB110_Interf_Program_M1".Signals_ExPlant[1].shot_end,
           OUT_ServiceShot          := "DB110_Interf_Program_M1".Signals_ExPlant[1].Service_mode,
           IO_Status                := "DB110_Interf_Program_M1".Status_ExPlant[1],
           IO_Fault                 := "DB825_Error_Interface".Interface_externalPlant[1],
           IO_NewFault              := "DB009_Faults".Faultschanging_M1,
           IO_FaultLevel_1          := "DB009_Faults".Faults_FKT_Grp_1_M1,
           IO_FaultLevel_2          := "DB009_Faults".Faults_FKT_Grp_2_M1,
           IO_FaultLevel_3          := "DB009_Faults".Faults_FKT_Grp_3_M1
         );
   //-----

   NoInterfaceMH1:NOP   0;
END_REGION

REGION Network 3: Send Process datas to KMI
         JU    M02c;

         A     "DB619_State_MPart".Operationmode[1].Auto;
         A     "DB704_MH_Value".Mixinghead[1].Conf_IntWithPlantInerface;
         CLR;
         JC    M02c;

         AN    "DB619_State_MPart".Cycle[1].PulsShotend;
         JC    M030;

         L     "DB919_ShotResultMach".ShotResult_Ma[1].General.MH_No;
         T     "DB149_KMI_FRA_Data".Measured_values_to_INT01.MH_Number;

   M030: NOP   0;

   // Flag shotend  (200ms)
   //    U     "DB149_KMI_FRA_Data".Signals_INT01.PU_Shot_End
         O     "DB005_RS<->Extern".MC_Interface[1].Data_to_MC.Shot_end;
         O     "DB005_RS<->Extern".MC_Interface[2].Data_to_MC.Shot_end;
         O     "DB005_RS<->Extern".MC_Interface[3].Data_to_MC.Shot_end;
         O     "DB005_RS<->Extern".MC_Interface[4].Data_to_MC.Shot_end;
         L     S5T#200MS;
         SE    "T_Delay_Send_Data_KMI";

         A     "T_Delay_Send_Data_KMI";
         FN    "Helpflag_Send_Data_KMI";
         =     "Send_Data_to_KMI";

         A     "Send_Data_to_KMI";
         =     "DB149_KMI_FRA_Data".Measured_values_to_INT01.Strobe_ProcessData;

   // Werte an FRA
   //-----------------------------------------------------------
         A     "DB149_KMI_FRA_Data".Measured_values_to_INT01.Strobe_ProcessData;
         JCN   M02d;
   ///
         L     "DB149_KMI_FRA_Data".Measured_values_to_INT01.MH_Number;
         T     "MH_Number_to_KMI":P;

         L     "DB919_ShotResultMach".ShotResult_Ma[1].General.PartWeight;
         L     10.0;
         *R;
         RND;
         T     "DB149_KMI_FRA_Data".Measured_values_to_INT01.Shot_Weight;
         T     "Shotwight_to_KMI":P;
   ///
         L     "DB919_ShotResultMach".ShotResult_Ma[1].General.FoamingTime;
         L     100.0;
         *R;
         RND;
         T     "DB149_KMI_FRA_Data".Measured_values_to_INT01.Shot_Time;
         T     "Shottime_to_KMI":P;

         L     "DB919_ShotResultMach".ShotResult_Ma[1].Component.Comp[1].TemperatureMH;
         L     10.0;
         *R;
         RND;
         T     "DB149_KMI_FRA_Data".Measured_values_to_INT01.Temperature_Poly;
         T     "Temp_C1_MH_to_KMI":P;
   ///
         L     "DB919_ShotResultMach".ShotResult_Ma[1].Component.Comp[2].TemperatureMH;
         L     10.0;
         *R;
         RND;
         T     "DB149_KMI_FRA_Data".Measured_values_to_INT01.Temperature_Iso;
         T     "Temp_C2_MH_to_KMI":P;

   ///
         L     "DB919_ShotResultMach".ShotResult_Ma[1].Component.Comp[1].Mixingratio;
         L     10.0;
         *R;
         RND;
         T     "DB149_KMI_FRA_Data".Measured_values_to_INT01.Mix_Rate_Poly;
         T     "Ratio_C1_to_KMI":P;

   ///
         L     "DB919_ShotResultMach".ShotResult_Ma[1].Component.Comp[2].Mixingratio;
         L     10.0;
         *R;
         RND;
         T     "DB149_KMI_FRA_Data".Measured_values_to_INT01.Mix_Rate_Iso;
         T     "Ratio_C2_to_KMI":P;
   ///
         L     "DB919_ShotResultMach".ShotResult_Ma[1].Component.Comp[1].PressureMH;
         L     10.0;
         *R;
         RND;
         T     "DB149_KMI_FRA_Data".Measured_values_to_INT01.Pressure_Poly;
         T     "Pressure_C1_MH_to_KMI":P;
   ///
         L     "DB919_ShotResultMach".ShotResult_Ma[1].Component.Comp[2].PressureMH;
         L     10.0;
         *R;
         RND;
         T     "DB149_KMI_FRA_Data".Measured_values_to_INT01.Pressure_Iso;
         T     "Pressure_C2_MH_to_KMI":P;

   // Alarmbits an FRA
   M02d: A     "DB009_Faults".Faults_Reset_FKT_M1;
         R     "DB149_KMI_FRA_Data".Measured_values_to_INT01.Alarm_flow_K1;
         R     "DB149_KMI_FRA_Data".Measured_values_to_INT01.Alarm_flow_K2;
         R     "DB149_KMI_FRA_Data".Measured_values_to_INT01.Alarm_press_K1;
         R     "DB149_KMI_FRA_Data".Measured_values_to_INT01.Alarm_press_K2;
         R     "DB149_KMI_FRA_Data".Measured_values_to_INT01.Alarm_temp_K1;
         R     "DB149_KMI_FRA_Data".Measured_values_to_INT01.Alarm_temp_K2;
         R     "DB149_KMI_FRA_Data".Measured_values_to_INT01.Alarm_shottime;

         A     "DB110_Interf_Program_M1".Status_ExPlant[1].IF_is_selected;
         JCN   Ala1;

         O     "DB823_Error_Metering".Flow_Component[1].Alarm_limit_plus;
         O     "DB823_Error_Metering".Flow_Component[1].Alarm_limit_minus;
         S     "DB149_KMI_FRA_Data".Measured_values_to_INT01.Alarm_flow_K1;

         O     "DB823_Error_Metering".Flow_Component[2].Alarm_limit_plus;
         O     "DB823_Error_Metering".Flow_Component[2].Alarm_limit_minus;
         S     "DB149_KMI_FRA_Data".Measured_values_to_INT01.Alarm_flow_K2;

         O     "DB824_Error_MH_CP".Pressure[1, 1].Alarm_limit_plus;
         O     "DB824_Error_MH_CP".Pressure[1, 1].Alarm_limit_minus;
         S     "DB149_KMI_FRA_Data".Measured_values_to_INT01.Alarm_press_K1;

         O     "DB824_Error_MH_CP".Pressure[2, 1].Alarm_limit_plus;
         O     "DB824_Error_MH_CP".Pressure[2, 1].Alarm_limit_minus;
         S     "DB149_KMI_FRA_Data".Measured_values_to_INT01.Alarm_press_K2;

         O     "DB824_Error_MH_CP".Temperature[1, 1].Alarm_limit_plus;
         O     "DB824_Error_MH_CP".Temperature[1, 1].Alarm_limit_minus;
         S     "DB149_KMI_FRA_Data".Measured_values_to_INT01.Alarm_temp_K1;

         O     "DB824_Error_MH_CP".Temperature[2, 1].Alarm_limit_plus;
         O     "DB824_Error_MH_CP".Temperature[2, 1].Alarm_limit_minus;
         S     "DB149_KMI_FRA_Data".Measured_values_to_INT01.Alarm_temp_K2;

         O     "DB829_Error_Machine".Foaming_Time[1].Alarm_limit_plus;
         O     "DB829_Error_Machine".Foaming_Time[1].Alarm_limit_minus;
         S     "DB149_KMI_FRA_Data".Measured_values_to_INT01.Alarm_shottime;

   Ala1: NOP   0;

   // Datas to Int Alarmbits
         L     %DB149.DBW38;
         T     "Alarm_Bits_to_KMI":P;

   M02c: NOP   0;
END_REGION

REGION Network 4: Release foaming interface mouldcarrier
END_REGION

REGION Network 5: Signals foaming a tool (mould)
   //----
         ON    "DB619_State_MPart".Cycle[1].running;
         O(;
         A     "DB619_State_MPart".Cycle[1].LastStanbyTimeTool;
         AN    "DB619_State_MPart".Cycle[1].StandByTimeRuns;
         );
         R     "DB619_State_MPart".Cycle[1].LastShotinToolFinished;
   //---
         A     "DB619_State_MPart".ToolMa[1].StationFinished;
         A     "DB619_State_MPart".Cycle[1].running;
         AN    "DB619_State_MPart".Cycle[1].LastShotinToolFinished;
         S     "DB619_State_MPart".Cycle[1].LastShotinTool;
   //---
         O(;
         A     "DB110_Interf_Program_M1".Bits.LastShotAtThisMachine;
         A     "DB619_State_MPart".Cycle[1].Pulse_ToolFinished;
         );
         O(;
         AN    "DB619_State_MPart".ToolMa[1].ShotFound;
         A     "DB110_Interf_Program_M1".Bits.PulseShotEnd;
         );
         A     "DB619_State_MPart".Cycle[1].LastShotinTool;
         =     "DB110_Interf_Program_M1".Bits.PulseToolFinished;

         O     "DB110_Interf_Program_M1".Bits.PulseToolFinished;
         O     "DB619_State_MPart".Cycle[1].PulseCycleEnd;
         O(;
   //      U     "DB619_State_MPart".Cycle[1].PulsShotend
         A     "DB619_State_MPart".Cycle[1].LastShotinTool;
         );
         O(;
         AN    "DB619_State_MPart".Cycle[1].running;
         A     "DB619_State_MPart".Cycle[1].LastShotinTool;
         );
         FP    "DB110_Interf_Program_M1".Bits.HF_FP_PulseToolFinished;
         =     "DB619_State_MPart".Cycle[1].Pulse_ToolFinished;
         R     "DB619_State_MPart".Cycle[1].LastShotinTool;
         S     "DB619_State_MPart".Cycle[1].LastShotinToolFinished;

         A     "DB619_State_MPart".Cycle[1].LastShotinToolFinished;
         A     "DB619_State_MPart".Cycle[1].StandByTimeRuns;
         =     "DB619_State_MPart".Cycle[1].LastStanbyTimeTool;
         R     "DB619_State_MPart".Cycle[1].LastShotinTool;

         AN    "DB619_State_MPart".Cycle[1].Pulse_ToolFinished;
         JC    nw4e;
         L     "DB619_State_MPart".ToolMa[1].WorkCounter;
         L     1;
         +D;
         T     "DB619_State_MPart".ToolMa[1].WorkCounter;
   nw4e: NOP   0;
   //----
         A     "DB619_State_MPart".Cycle[1].running;
         R     "DB110_Interf_Program_M1".Bits.LastShotAtThisMachine;

         A     "DB619_State_MPart".Cycle[1].LastShotinTool;
         A     "DB619_State_MPart".ToolMa[1].ShotFound;
         S     "DB110_Interf_Program_M1".Bits.LastShotAtThisMachine;

         A     "DB619_State_MPart".Cycle[1].PulsShotend;
         =     "DB110_Interf_Program_M1".Bits.PulseShotEnd;

   //-----------------------------------------------------------------------------
   // Stop Interface if mould is not released
   //-----------------------------------------------------------------------------
         A     "DB619_State_MPart".ToolMa[1].StationFinished;
         AN    "DB619_State_MPart".Cycle[1].running;
         FP    "DB110_Interf_Program_M1".Bits.HF_FP_MouldNotReleased;
         =     "DB110_Interf_Program_M1".Bits.MouldNotReleased;